// TIA Portal project "Liikennevalot" (V16)

(* hardware
DEVICE "S7-1200 station_1"  S7-1200 Station
   slot 0: "Rack_0"  S7-1200 Rack  Rack  V1.0
   slot 1: "PLC_1"  CPU 1215C DC/DC/DC  6ES7 215-1AG40-0XB0  V4.4
DEVICE "HMI_1"  KTP1200 Basic PN
   slot 0: "HMI_1"  KTP1200 Basic PN  6AV2 123-2MB03-0AX0  16.0.0.0
   slot 1: "HMI_RT_1"  KTP1200 Basic PN  6AV2 123-2MB03-0AX0  16.0.0.0
   slot 5: "HMI_1.IE_CP_1"  PROFINET Interface  16.0.0.0
      slot 1: "PROFINET Interface_1"  PROFINET Interface
         slot 1: "Port_1"  Port
*)

// ===== PLC "PLC_1"  CPU 1215C DC/DC/DC =====

VAR_GLOBAL   // PLC tag table "Default tag table"
   "Car_Yellow" AT %Q0.0 : Bool;
   "Car_Red" AT %Q0.1 : Bool;
   "Car_Green" AT %Q0.2 : Bool;
   "Pedestrian_Red" AT %Q0.3 : Bool;
   "Pedestrian_Green" AT %Q0.4 : Bool;
   "Pedestrian_Yellow" AT %Q0.5 : Bool;
   "Pedestrian_Button" AT %M0.0 : Bool;
   "Memory1" AT %Q0.6 : Bool;
   "Memory2" AT %Q0.7 : Bool;
END_VAR

// folder: System blocks/Program resources

DATA_BLOCK "Timer_1"   // DB1
{ S7_Optimized_Access := 'TRUE' }
AUTHOR : Simatic
FAMILY : IEC
NAME : IEC_TMR
VERSION : 1.0
// stored: InstanceOfName IEC_TIMER
"IEC_TIMER"
BEGIN
END_DATA_BLOCK

DATA_BLOCK "Timer_2"   // DB2
{ S7_Optimized_Access := 'TRUE' }
AUTHOR : Simatic
FAMILY : IEC
NAME : IEC_TMR
VERSION : 1.0
// stored: InstanceOfName IEC_TIMER
"IEC_TIMER"
BEGIN
END_DATA_BLOCK

DATA_BLOCK "Timer_3"   // DB3
{ S7_Optimized_Access := 'TRUE' }
AUTHOR : Simatic
FAMILY : IEC
NAME : IEC_TMR
VERSION : 1.0
// stored: InstanceOfName IEC_TIMER
"IEC_TIMER"
BEGIN
END_DATA_BLOCK

// folder: (top level)

ORGANIZATION_BLOCK "Main"   // OB1, FBD, ProgramCycle
TITLE = "Main Program Sweep (Cycle)"
{ S7_Optimized_Access := 'TRUE' }
VERSION : 0.1
   VAR_INPUT
      Initial_Call : Bool;   // Initial call of this OB
      Remanence : Bool;   // =True, if remanent data are available
   END_VAR
   VAR_TEMP   // added for the SCL form of the ladder/FBD networks
      _w1 : Bool;
   END_VAR
BEGIN

REGION Network 1
   // Traffic lights for cars
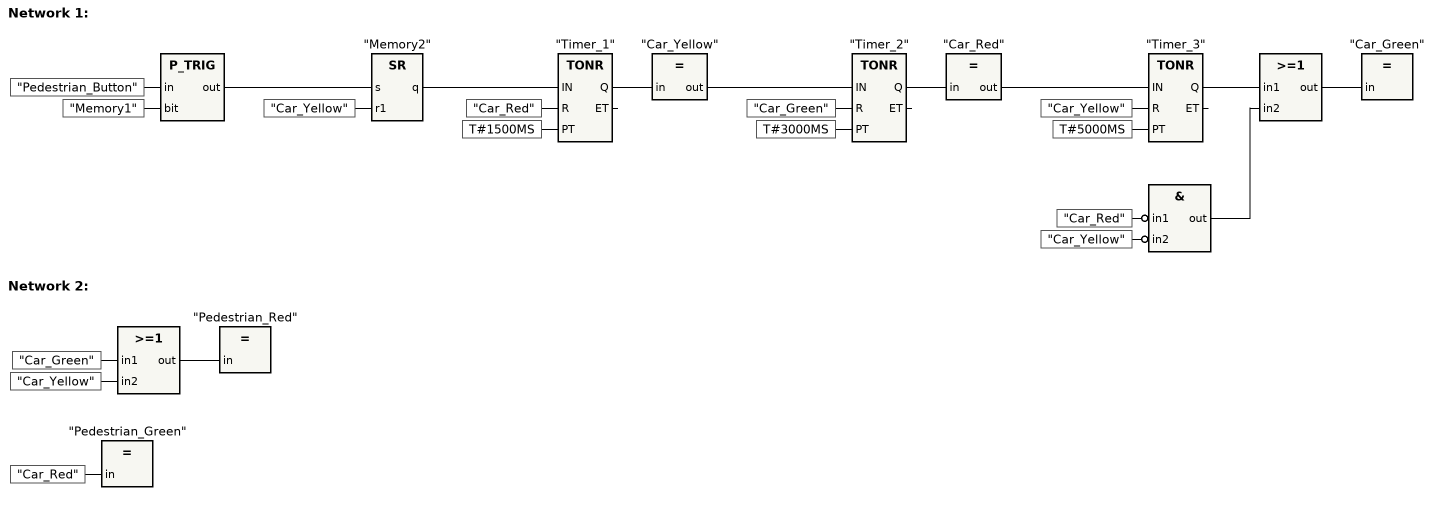
   #_w1 := "Pedestrian_Button" AND NOT "Memory1";   // rising edge
   "Memory1" := "Pedestrian_Button";
   IF #_w1 THEN
       "Memory2" := TRUE;   // SR flip-flop
   END_IF;
   IF "Car_Yellow" THEN "Memory2" := FALSE; END_IF;
   "Timer_1".TONR(IN := "Memory2", R := "Car_Red", PT := T#1500MS);
   "Car_Yellow" := "Timer_1".Q;
   "Timer_2".TONR(IN := "Timer_1".Q, R := "Car_Green", PT := T#3000MS);
   "Car_Red" := "Timer_2".Q;
   "Timer_3".TONR(IN := "Timer_2".Q, R := "Car_Yellow", PT := T#5000MS);
   "Car_Green" := "Timer_3".Q OR (NOT "Car_Red" AND NOT "Car_Yellow");
END_REGION

REGION Network 2
   // Traffic lights for pedestrians
   "Pedestrian_Red" := "Car_Green" OR "Car_Yellow";
   "Pedestrian_Green" := "Car_Red";
END_REGION
END_ORGANIZATION_BLOCK

(* ===== HMI "HMI_RT_1" =====
system functions are stored by id; their names below are inferred from use
connection "HMI_Connection_1": ETHERNET, SMART_S7_1200_OMS

HMI tags "Default tag table"
   "Tag_ScreenNumber" : UInt AT %DB1.DBW0
   "Car_Red" : Bool = PLC Car_Red AT %Q0.1, 1 s
   "Car_Green" : Bool = PLC Car_Green AT %Q0.2, 1 s
   "Car_Yellow" : Bool = PLC Car_Yellow AT %Q0.0, 1 s
   "Pedesterian_Green" : Bool = PLC Pedestrian_Green AT %Q0.4, 1 s
   "Pedestrian_Red" : Bool = PLC Pedestrian_Red AT %Q0.3, 1 s
   "Pedestrian_Button" : Bool AT %M0.0, 1 s

Template "Template_1" 1280x800
   SymbolicIOField "Symbolic_IO_Field_Screen" at 87,9 size 1086x30; TextOff '0'; TextOn '1'; TextList "TextList_ScreenNames"
      ProcessValue <- "Tag_ScreenNumber"
      on Change: ActivateScreenByNumber("Tag_ScreenNumber", 0)
   DateTimeField "HmiScreenItemData" at 1175,24 size 105x24
   DateTimeField "HmiScreenItemData_1" at 1175,0 size 105x24
   GraphicView "Logo" at 0,0 size 85x48; Picture "Logo of HMI_1"

screen "Root screen" 1280x800, template "Template_1"
   on GenerateScreen: SetTag("Pedestrian_Button", 1)
   Circle "Circle_1" at 80,92 size 89x89
      Appearance <- "Pedestrian_Red"
   Circle "Circle_2" at 80,191 size 89x89
      Appearance <- "Pedesterian_Green"
   Button "Button_1" at 80,437 size 96x32; TextOff 'Text'
      on Press: function_b14e0dd5("Pedestrian_Button", 0)
      Appearance <- "Pedestrian_Button"
   Circle "Circle_4" at 964,92 size 89x89
      Appearance <- "Car_Red"
   Circle "Circle_5" at 964,191 size 89x89
      Appearance <- "Car_Yellow"
   Circle "Circle_6" at 964,290 size 89x89
      Appearance <- "Car_Green"
   TextField "Text field_1" at 964,412 size 183x25; Text 'Traffic lights for cars'
   TextField "Text field_2" at 80,404 size 248x25; Text 'Traffic lights for pedestrians'
*)